REGION Network 2: Auto Initiated = Set Step to 1
   // Once the pulse has expired, with the system still in automatic, the step is set to 1
   RUNG wire#powerrail
      { S7_Templates := "SrcType := Int" } EQ_Contact(in1 := #CRNT_STEP, in2 := 0)
      I_Contact( #RST )
      Move(in := 1, out1 => #CRNT_STEP)
   END_RUNG
   // the same network as SCL:
   IF (#CRNT_STEP = 0) AND NOT #RST THEN #CRNT_STEP := 1; END_IF;
END_REGION

REGION Network 3: Sequence Running
   // Determination that the sequence is running
   RUNG wire#powerrail
      { S7_Templates := "SrcType := Int" } NE_Contact(in1 := #CRNT_STEP, in2 := 0)
      Coil( #RNG )
   END_RUNG
   // the same network as SCL:
   #RNG := #CRNT_STEP <> 0;
END_REGION

REGION Network 4: Step 001 = Confirm Auto Conditions Ok
   // Requires all conditions for auto ok to proceed
   RUNG wire#powerrail
      #STEP_001(SN := 1, CS := #CRNT_STEP, MST := "86_Times".STEP_MAX_TIME_STP_001, SC :=, BPFLT := true, AMST :=, FLT :=, ACT =>, DN =>)
      Contact( #STEP_001.DN )
      Move(in := 5, out1 => #CRNT_STEP)
   END_RUNG
   // the same network as SCL:
   #STEP_001(SN := 1, CS := #CRNT_STEP, MST := "86_Times".STEP_MAX_TIME_STP_001, BPFLT := true, ENO => #_w1);   // "500_SEQ_STEP"
   IF #_w1 AND #STEP_001.DN THEN #CRNT_STEP := 5; END_IF;
END_REGION

REGION Network 5: Step 005 = Wait For BWTS In Pre-Dwell or Dwell & ReOx
   // BWTS Active throughout
   RUNG wire#powerrail
      #STEP_005(SN := 5, CS := #CRNT_STEP, MST := "86_Times".STEP_MAX_TIME_STP_005, SC :=, BPFLT := true, AMST :=, FLT :=, ACT =>, DN =>)
      Contact( #STEP_005.DN )
      Move(in := 10, out1 => #CRNT_STEP)
   END_RUNG
   // the same network as SCL:
   #STEP_005(SN := 5, CS := #CRNT_STEP, MST := "86_Times".STEP_MAX_TIME_STP_005, BPFLT := true, ENO => #_w1);   // "500_SEQ_STEP"
   IF #_w1 AND #STEP_005.DN THEN #CRNT_STEP := 10; END_IF;
END_REGION

REGION Network 6: Step 010 = Wait For Prepare Gas Command (DeOx = Step 20, ReOx = Step 40)
   // BWTS Sends prepare gas command an hour prior to physical requirement
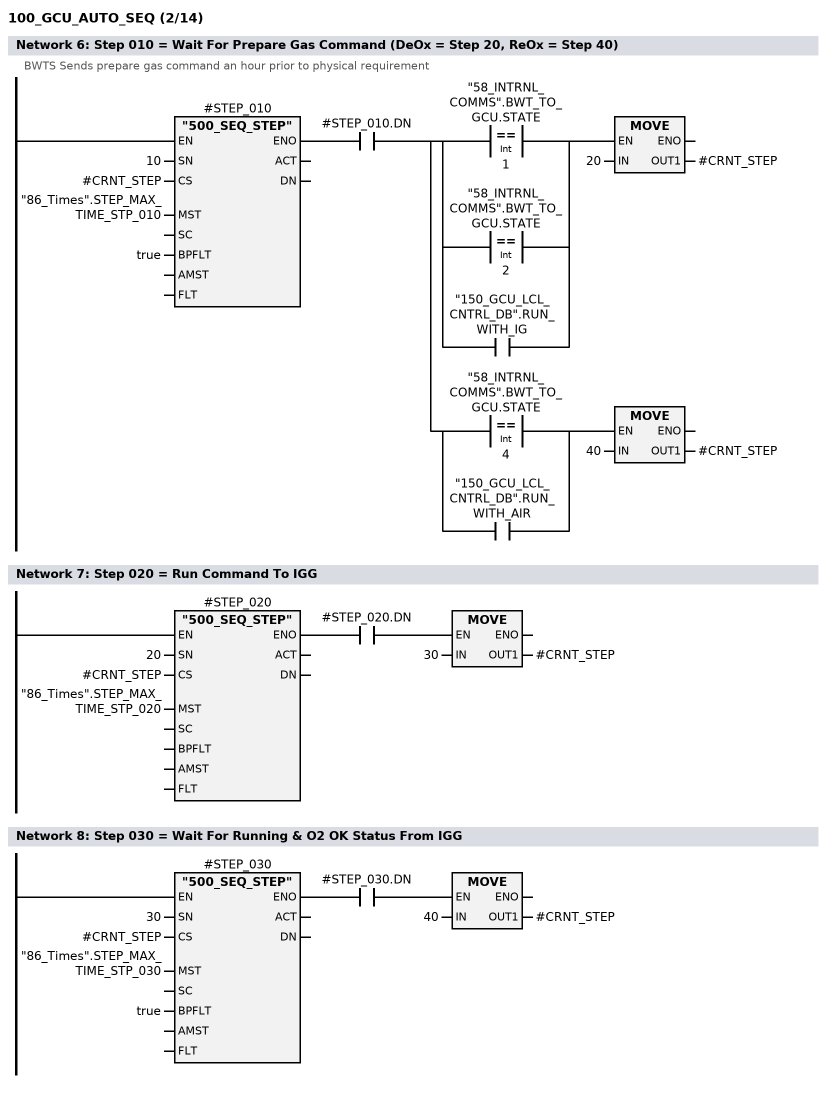
   RUNG wire#powerrail
      #STEP_010(SN := 10, CS := #CRNT_STEP, MST := "86_Times".STEP_MAX_TIME_STP_010, SC :=, BPFLT := true, AMST :=, FLT :=, ACT =>, DN =>)
      Contact( #STEP_010.DN )
      wire#w1
      { S7_Templates := "SrcType := Int" } EQ_Contact(in1 := "58_INTRNL_COMMS".BWT_TO_GCU.STATE, in2 := 1)
      wire#w2
      Move(in := 20, out1 => #CRNT_STEP)
   END_RUNG
   RUNG wire#w1
      { S7_Templates := "SrcType := Int" } EQ_Contact(in1 := "58_INTRNL_COMMS".BWT_TO_GCU.STATE, in2 := 2)
   END_RUNG wire#w2
   RUNG wire#w1
      Contact( "150_GCU_LCL_CNTRL_DB".RUN_WITH_IG )
   END_RUNG wire#w2
   RUNG wire#w1
      { S7_Templates := "SrcType := Int" } EQ_Contact(in1 := "58_INTRNL_COMMS".BWT_TO_GCU.STATE, in2 := 4)
      wire#w3
      Move(in := 40, out1 => #CRNT_STEP)
   END_RUNG
   RUNG wire#w1
      Contact( "150_GCU_LCL_CNTRL_DB".RUN_WITH_AIR )
   END_RUNG wire#w3
   // the same network as SCL:
   #STEP_010(SN := 10, CS := #CRNT_STEP, MST := "86_Times".STEP_MAX_TIME_STP_010, BPFLT := true, ENO => #_w1);   // "500_SEQ_STEP"
   #_w2 := #_w1 AND #STEP_010.DN;
   IF #_w2 AND (("58_INTRNL_COMMS".BWT_TO_GCU.STATE = 1) OR ("58_INTRNL_COMMS".BWT_TO_GCU.STATE = 2) OR "150_GCU_LCL_CNTRL_DB".RUN_WITH_IG) THEN
       #CRNT_STEP := 20;
   END_IF;
   IF #_w2 AND (("58_INTRNL_COMMS".BWT_TO_GCU.STATE = 4) OR "150_GCU_LCL_CNTRL_DB".RUN_WITH_AIR) THEN
       #CRNT_STEP := 40;
   END_IF;
END_REGION

REGION Network 7: Step 020 = Run Command To IGG
   RUNG wire#powerrail
      #STEP_020(SN := 20, CS := #CRNT_STEP, MST := "86_Times".STEP_MAX_TIME_STP_020, SC :=, BPFLT :=, AMST :=, FLT :=, ACT =>, DN =>)
      Contact( #STEP_020.DN )
      Move(in := 30, out1 => #CRNT_STEP)
   END_RUNG
   // the same network as SCL:
   #STEP_020(SN := 20, CS := #CRNT_STEP, MST := "86_Times".STEP_MAX_TIME_STP_020, ENO => #_w1);   // "500_SEQ_STEP"
   IF #_w1 AND #STEP_020.DN THEN #CRNT_STEP := 30; END_IF;
END_REGION

REGION Network 8: Step 030 = Wait For Running & O2 OK Status From IGG
   RUNG wire#powerrail
      #STEP_030(SN := 30, CS := #CRNT_STEP, MST := "86_Times".STEP_MAX_TIME_STP_030, SC :=, BPFLT := true, AMST :=, FLT :=, ACT =>, DN =>)
      Contact( #STEP_030.DN )
      Move(in := 40, out1 => #CRNT_STEP)
   END_RUNG
   // the same network as SCL:
   #STEP_030(SN := 30, CS := #CRNT_STEP, MST := "86_Times".STEP_MAX_TIME_STP_030, BPFLT := true, ENO => #_w1);   // "500_SEQ_STEP"
   IF #_w1 AND #STEP_030.DN THEN #CRNT_STEP := 40; END_IF;
END_REGION

REGION Network 9: Step 040 = Wait For Supply Gas Command
   // Gas available status to BWTS
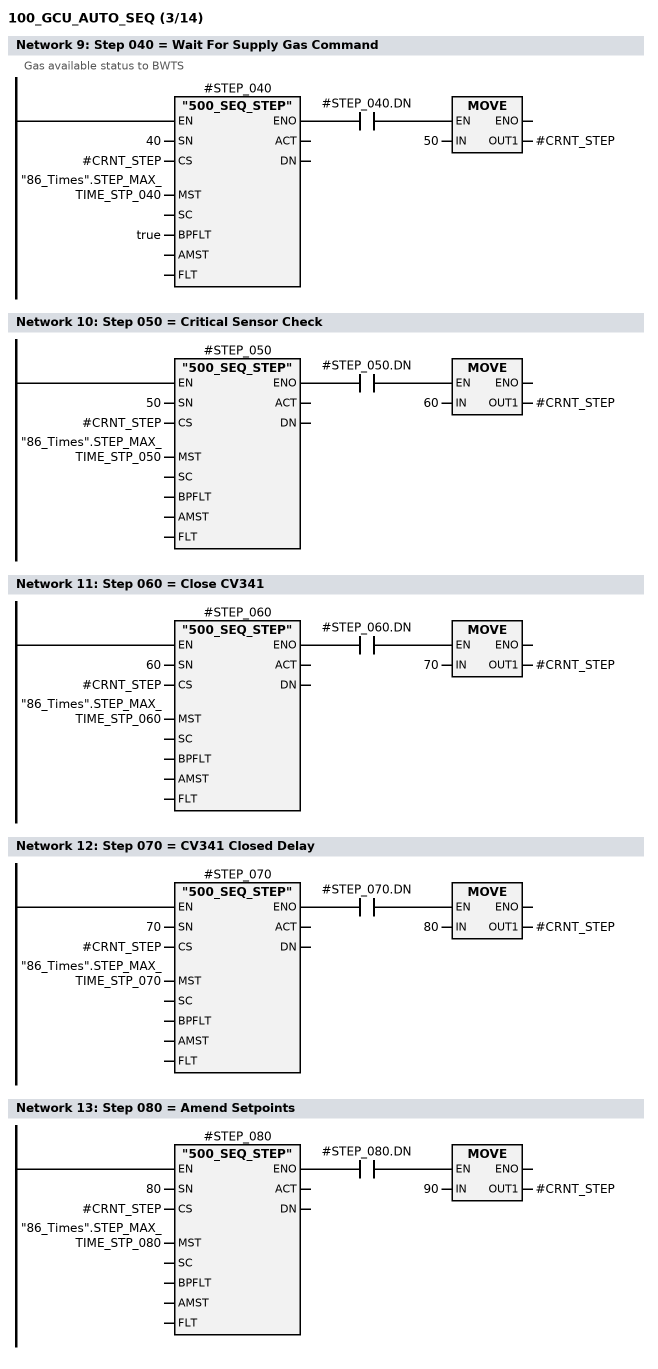
   RUNG wire#powerrail
      #STEP_040(SN := 40, CS := #CRNT_STEP, MST := "86_Times".STEP_MAX_TIME_STP_040, SC :=, BPFLT := true, AMST :=, FLT :=, ACT =>, DN =>)
      Contact( #STEP_040.DN )
      Move(in := 50, out1 => #CRNT_STEP)
   END_RUNG
   // the same network as SCL:
   #STEP_040(SN := 40, CS := #CRNT_STEP, MST := "86_Times".STEP_MAX_TIME_STP_040, BPFLT := true, ENO => #_w1);   // "500_SEQ_STEP"
   IF #_w1 AND #STEP_040.DN THEN #CRNT_STEP := 50; END_IF;
END_REGION

REGION Network 10: Step 050 = Critical Sensor Check
   RUNG wire#powerrail
      #STEP_050(SN := 50, CS := #CRNT_STEP, MST := "86_Times".STEP_MAX_TIME_STP_050, SC :=, BPFLT :=, AMST :=, FLT :=, ACT =>, DN =>)
      Contact( #STEP_050.DN )
      Move(in := 60, out1 => #CRNT_STEP)
   END_RUNG
   // the same network as SCL:
   #STEP_050(SN := 50, CS := #CRNT_STEP, MST := "86_Times".STEP_MAX_TIME_STP_050, ENO => #_w1);   // "500_SEQ_STEP"
   IF #_w1 AND #STEP_050.DN THEN #CRNT_STEP := 60; END_IF;
END_REGION

REGION Network 11: Step 060 = Close CV341
   RUNG wire#powerrail
      #STEP_060(SN := 60, CS := #CRNT_STEP, MST := "86_Times".STEP_MAX_TIME_STP_060, SC :=, BPFLT :=, AMST :=, FLT :=, ACT =>, DN =>)
      Contact( #STEP_060.DN )
      Move(in := 70, out1 => #CRNT_STEP)
   END_RUNG
   // the same network as SCL:
   #STEP_060(SN := 60, CS := #CRNT_STEP, MST := "86_Times".STEP_MAX_TIME_STP_060, ENO => #_w1);   // "500_SEQ_STEP"
   IF #_w1 AND #STEP_060.DN THEN #CRNT_STEP := 70; END_IF;
END_REGION

REGION Network 12: Step 070 = CV341 Closed Delay
   RUNG wire#powerrail
      #STEP_070(SN := 70, CS := #CRNT_STEP, MST := "86_Times".STEP_MAX_TIME_STP_070, SC :=, BPFLT :=, AMST :=, FLT :=, ACT =>, DN =>)
      Contact( #STEP_070.DN )
      Move(in := 80, out1 => #CRNT_STEP)
   END_RUNG
   // the same network as SCL:
   #STEP_070(SN := 70, CS := #CRNT_STEP, MST := "86_Times".STEP_MAX_TIME_STP_070, ENO => #_w1);   // "500_SEQ_STEP"
   IF #_w1 AND #STEP_070.DN THEN #CRNT_STEP := 80; END_IF;
END_REGION

REGION Network 13: Step 080 = Amend Setpoints
   RUNG wire#powerrail
      #STEP_080(SN := 80, CS := #CRNT_STEP, MST := "86_Times".STEP_MAX_TIME_STP_080, SC :=, BPFLT :=, AMST :=, FLT :=, ACT =>, DN =>)
      Contact( #STEP_080.DN )
      Move(in := 90, out1 => #CRNT_STEP)
   END_RUNG
   // the same network as SCL:
   #STEP_080(SN := 80, CS := #CRNT_STEP, MST := "86_Times".STEP_MAX_TIME_STP_080, ENO => #_w1);   // "500_SEQ_STEP"
   IF #_w1 AND #STEP_080.DN THEN #CRNT_STEP := 90; END_IF;
END_REGION

REGION Network 14: Step 090 = Open CV358
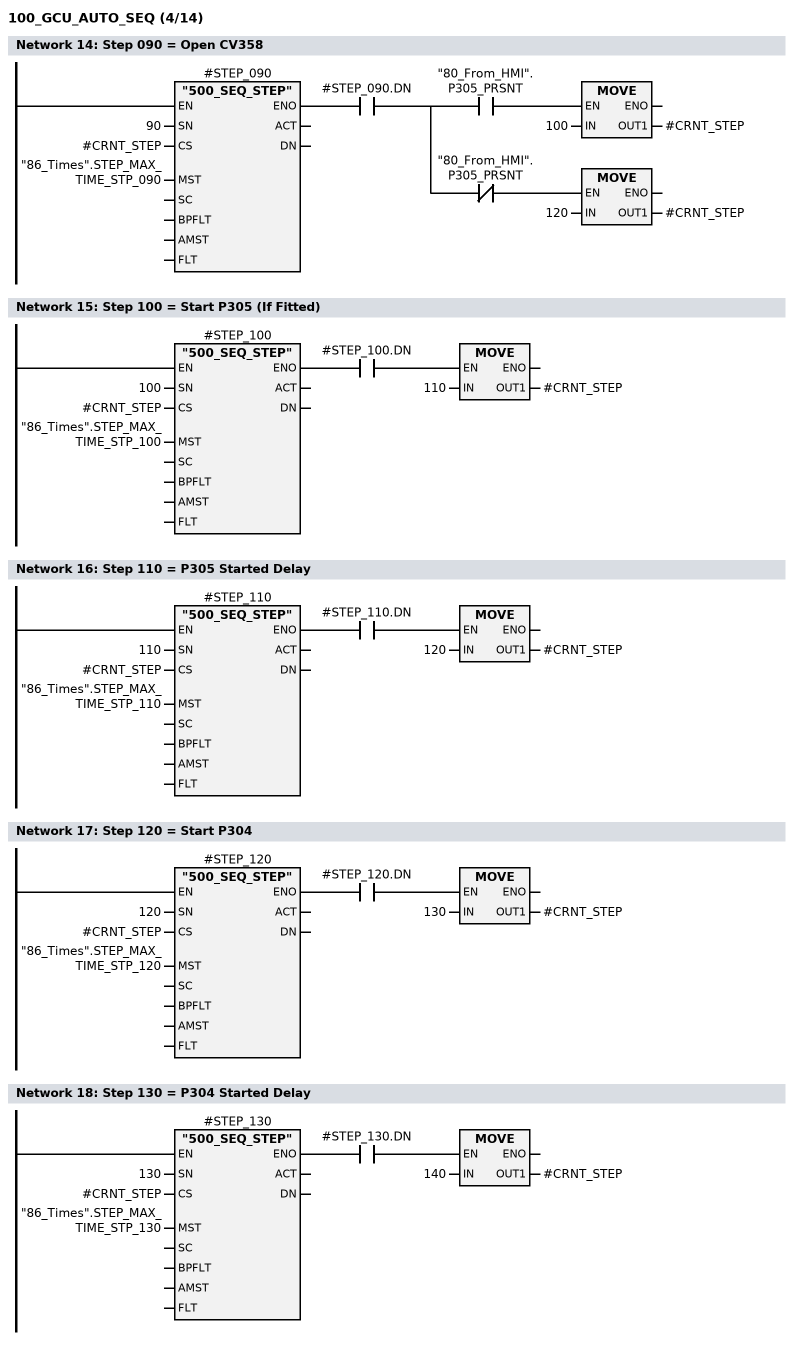
   RUNG wire#powerrail
      #STEP_090(SN := 90, CS := #CRNT_STEP, MST := "86_Times".STEP_MAX_TIME_STP_090, SC :=, BPFLT :=, AMST :=, FLT :=, ACT =>, DN =>)
      Contact( #STEP_090.DN )
      wire#w1
      Contact( "80_From_HMI".P305_PRSNT )
      Move(in := 100, out1 => #CRNT_STEP)
   END_RUNG
   RUNG wire#w1
      I_Contact( "80_From_HMI".P305_PRSNT )
      Move(in := 120, out1 => #CRNT_STEP)
   END_RUNG
   // the same network as SCL:
   #STEP_090(SN := 90, CS := #CRNT_STEP, MST := "86_Times".STEP_MAX_TIME_STP_090, ENO => #_w1);   // "500_SEQ_STEP"
   #_w2 := #_w1 AND #STEP_090.DN;
   IF #_w2 AND "80_From_HMI".P305_PRSNT THEN #CRNT_STEP := 100; END_IF;
   IF #_w2 AND NOT "80_From_HMI".P305_PRSNT THEN #CRNT_STEP := 120; END_IF;
END_REGION

REGION Network 15: Step 100 = Start P305 (If Fitted)
   RUNG wire#powerrail
      #STEP_100(SN := 100, CS := #CRNT_STEP, MST := "86_Times".STEP_MAX_TIME_STP_100, SC :=, BPFLT :=, AMST :=, FLT :=, ACT =>, DN =>)
      Contact( #STEP_100.DN )
      Move(in := 110, out1 => #CRNT_STEP)
   END_RUNG
   // the same network as SCL:
   #STEP_100(SN := 100, CS := #CRNT_STEP, MST := "86_Times".STEP_MAX_TIME_STP_100, ENO => #_w1);   // "500_SEQ_STEP"
   IF #_w1 AND #STEP_100.DN THEN #CRNT_STEP := 110; END_IF;
END_REGION

REGION Network 16: Step 110 = P305 Started Delay
   RUNG wire#powerrail
      #STEP_110(SN := 110, CS := #CRNT_STEP, MST := "86_Times".STEP_MAX_TIME_STP_110, SC :=, BPFLT :=, AMST :=, FLT :=, ACT =>, DN =>)
      Contact( #STEP_110.DN )
      Move(in := 120, out1 => #CRNT_STEP)
   END_RUNG
   // the same network as SCL:
   #STEP_110(SN := 110, CS := #CRNT_STEP, MST := "86_Times".STEP_MAX_TIME_STP_110, ENO => #_w1);   // "500_SEQ_STEP"
   IF #_w1 AND #STEP_110.DN THEN #CRNT_STEP := 120; END_IF;
END_REGION

REGION Network 17: Step 120 = Start P304
   RUNG wire#powerrail
      #STEP_120(SN := 120, CS := #CRNT_STEP, MST := "86_Times".STEP_MAX_TIME_STP_120, SC :=, BPFLT :=, AMST :=, FLT :=, ACT =>, DN =>)
      Contact( #STEP_120.DN )
      Move(in := 130, out1 => #CRNT_STEP)
   END_RUNG
   // the same network as SCL:
   #STEP_120(SN := 120, CS := #CRNT_STEP, MST := "86_Times".STEP_MAX_TIME_STP_120, ENO => #_w1);   // "500_SEQ_STEP"
   IF #_w1 AND #STEP_120.DN THEN #CRNT_STEP := 130; END_IF;
END_REGION

REGION Network 18: Step 130 = P304 Started Delay
   RUNG wire#powerrail
      #STEP_130(SN := 130, CS := #CRNT_STEP, MST := "86_Times".STEP_MAX_TIME_STP_130, SC :=, BPFLT :=, AMST :=, FLT :=, ACT =>, DN =>)
      Contact( #STEP_130.DN )
      Move(in := 140, out1 => #CRNT_STEP)
   END_RUNG
   // the same network as SCL:
   #STEP_130(SN := 130, CS := #CRNT_STEP, MST := "86_Times".STEP_MAX_TIME_STP_130, ENO => #_w1);   // "500_SEQ_STEP"
   IF #_w1 AND #STEP_130.DN THEN #CRNT_STEP := 140; END_IF;
END_REGION

REGION Network 19: Step 140 = GCU Tank Pre-Fill Delay
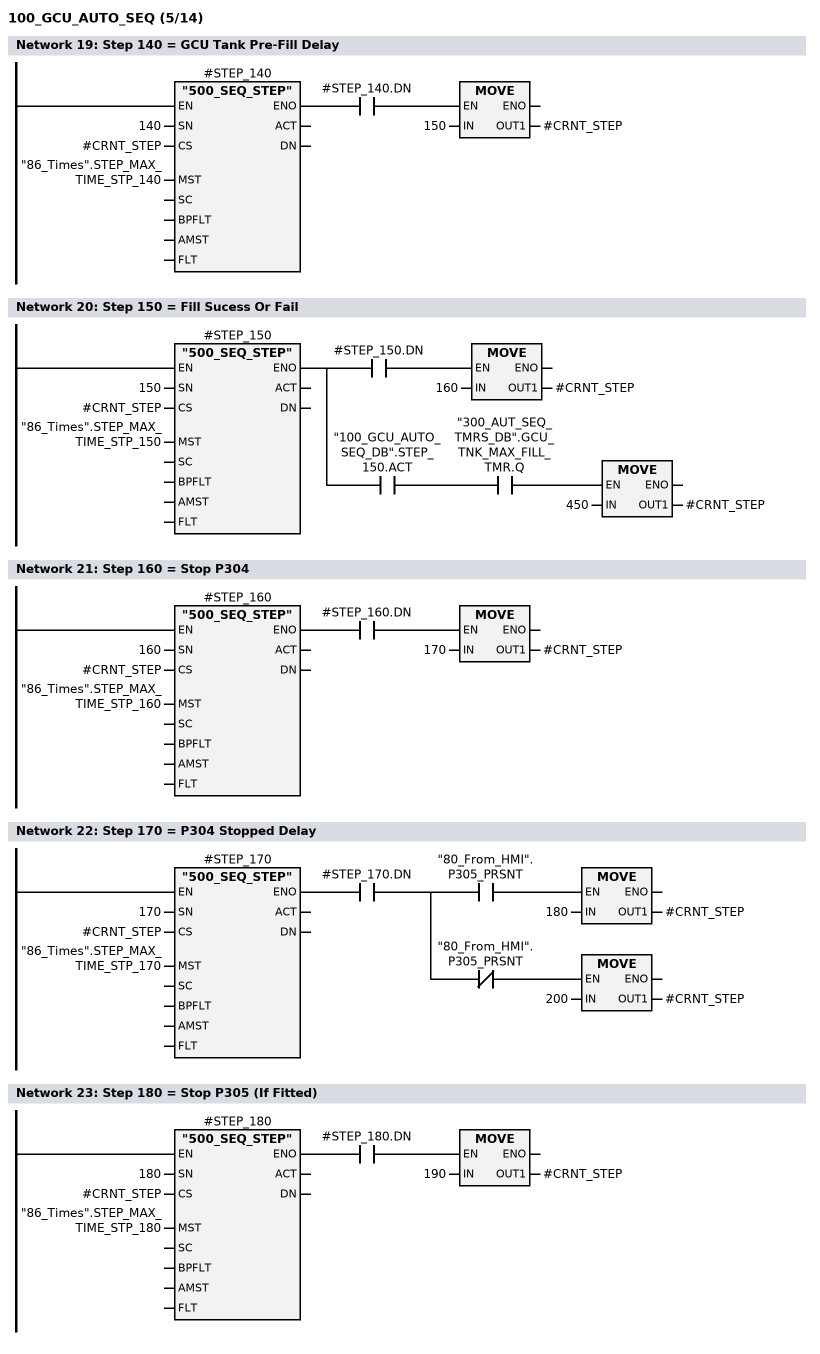
   RUNG wire#powerrail
      #STEP_140(SN := 140, CS := #CRNT_STEP, MST := "86_Times".STEP_MAX_TIME_STP_140, SC :=, BPFLT :=, AMST :=, FLT :=, ACT =>, DN =>)
      Contact( #STEP_140.DN )
      Move(in := 150, out1 => #CRNT_STEP)
   END_RUNG
   // the same network as SCL:
   #STEP_140(SN := 140, CS := #CRNT_STEP, MST := "86_Times".STEP_MAX_TIME_STP_140, ENO => #_w1);   // "500_SEQ_STEP"
   IF #_w1 AND #STEP_140.DN THEN #CRNT_STEP := 150; END_IF;
END_REGION

REGION Network 20: Step 150 = Fill Sucess Or Fail
   RUNG wire#powerrail
      #STEP_150(SN := 150, CS := #CRNT_STEP, MST := "86_Times".STEP_MAX_TIME_STP_150, SC :=, BPFLT :=, AMST :=, FLT :=, ACT =>, DN =>)
      wire#w1
      Contact( #STEP_150.DN )
      Move(in := 160, out1 => #CRNT_STEP)
   END_RUNG
   RUNG wire#w1
      Contact( "100_GCU_AUTO_SEQ_DB".STEP_150.ACT )
      Contact( "300_AUT_SEQ_TMRS_DB".GCU_TNK_MAX_FILL_TMR.Q )
      Move(in := 450, out1 => #CRNT_STEP)
   END_RUNG
   // the same network as SCL:
   #STEP_150(SN := 150, CS := #CRNT_STEP, MST := "86_Times".STEP_MAX_TIME_STP_150, ENO => #_w1);   // "500_SEQ_STEP"
   IF #_w1 AND #STEP_150.DN THEN #CRNT_STEP := 160; END_IF;
   IF #_w1 AND "100_GCU_AUTO_SEQ_DB".STEP_150.ACT AND "300_AUT_SEQ_TMRS_DB".GCU_TNK_MAX_FILL_TMR.Q THEN
       #CRNT_STEP := 450;
   END_IF;
END_REGION

REGION Network 21: Step 160 = Stop P304
   RUNG wire#powerrail
      #STEP_160(SN := 160, CS := #CRNT_STEP, MST := "86_Times".STEP_MAX_TIME_STP_160, SC :=, BPFLT :=, AMST :=, FLT :=, ACT =>, DN =>)
      Contact( #STEP_160.DN )
      Move(in := 170, out1 => #CRNT_STEP)
   END_RUNG
   // the same network as SCL:
   #STEP_160(SN := 160, CS := #CRNT_STEP, MST := "86_Times".STEP_MAX_TIME_STP_160, ENO => #_w1);   // "500_SEQ_STEP"
   IF #_w1 AND #STEP_160.DN THEN #CRNT_STEP := 170; END_IF;
END_REGION

REGION Network 22: Step 170 = P304 Stopped Delay
   RUNG wire#powerrail
      #STEP_170(SN := 170, CS := #CRNT_STEP, MST := "86_Times".STEP_MAX_TIME_STP_170, SC :=, BPFLT :=, AMST :=, FLT :=, ACT =>, DN =>)
      Contact( #STEP_170.DN )
      wire#w1
      Contact( "80_From_HMI".P305_PRSNT )
      Move(in := 180, out1 => #CRNT_STEP)
   END_RUNG
   RUNG wire#w1
      I_Contact( "80_From_HMI".P305_PRSNT )
      Move(in := 200, out1 => #CRNT_STEP)
   END_RUNG
   // the same network as SCL:
   #STEP_170(SN := 170, CS := #CRNT_STEP, MST := "86_Times".STEP_MAX_TIME_STP_170, ENO => #_w1);   // "500_SEQ_STEP"
   #_w2 := #_w1 AND #STEP_170.DN;
   IF #_w2 AND "80_From_HMI".P305_PRSNT THEN #CRNT_STEP := 180; END_IF;
   IF #_w2 AND NOT "80_From_HMI".P305_PRSNT THEN #CRNT_STEP := 200; END_IF;
END_REGION

REGION Network 23: Step 180 = Stop P305 (If Fitted)
   RUNG wire#powerrail
      #STEP_180(SN := 180, CS := #CRNT_STEP, MST := "86_Times".STEP_MAX_TIME_STP_180, SC :=, BPFLT :=, AMST :=, FLT :=, ACT =>, DN =>)
      Contact( #STEP_180.DN )
      Move(in := 190, out1 => #CRNT_STEP)
   END_RUNG
   // the same network as SCL:
   #STEP_180(SN := 180, CS := #CRNT_STEP, MST := "86_Times".STEP_MAX_TIME_STP_180, ENO => #_w1);   // "500_SEQ_STEP"
   IF #_w1 AND #STEP_180.DN THEN #CRNT_STEP := 190; END_IF;
END_REGION

REGION Network 24: Step 190 = P305 Stopped Delay
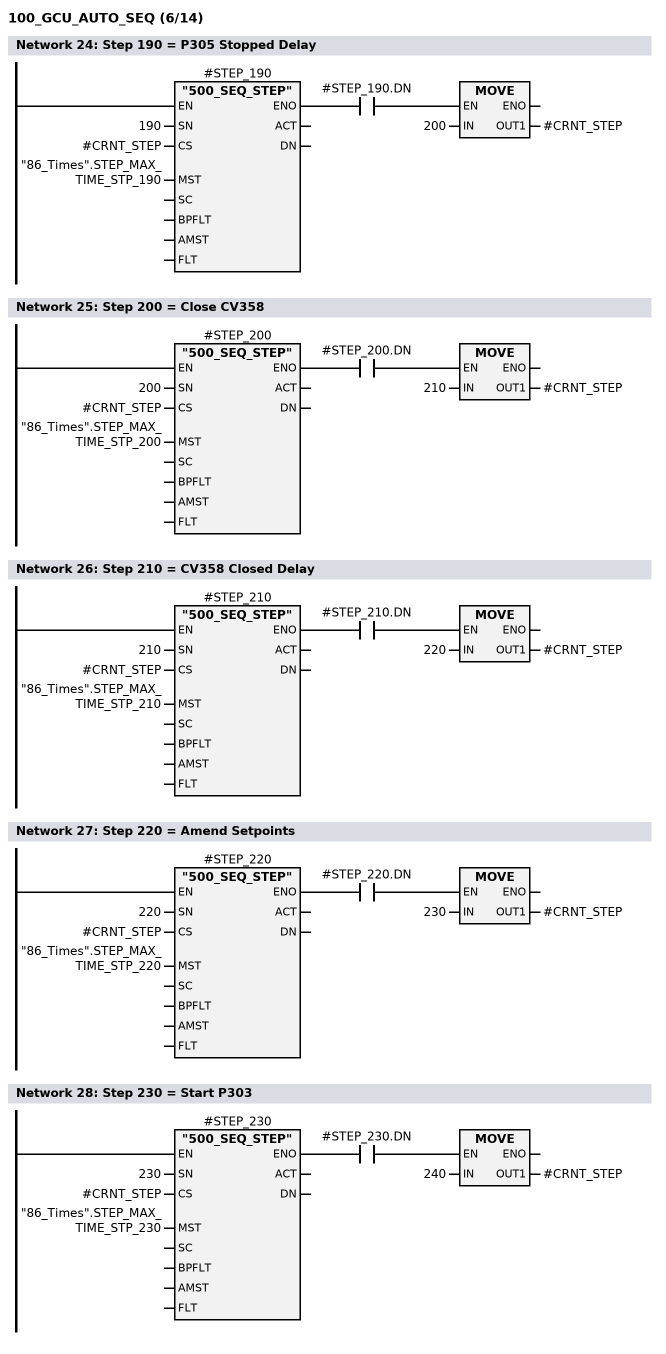
   RUNG wire#powerrail
      #STEP_190(SN := 190, CS := #CRNT_STEP, MST := "86_Times".STEP_MAX_TIME_STP_190, SC :=, BPFLT :=, AMST :=, FLT :=, ACT =>, DN =>)
      Contact( #STEP_190.DN )
      Move(in := 200, out1 => #CRNT_STEP)
   END_RUNG
   // the same network as SCL:
   #STEP_190(SN := 190, CS := #CRNT_STEP, MST := "86_Times".STEP_MAX_TIME_STP_190, ENO => #_w1);   // "500_SEQ_STEP"
   IF #_w1 AND #STEP_190.DN THEN #CRNT_STEP := 200; END_IF;
END_REGION

REGION Network 25: Step 200 = Close CV358
   RUNG wire#powerrail
      #STEP_200(SN := 200, CS := #CRNT_STEP, MST := "86_Times".STEP_MAX_TIME_STP_200, SC :=, BPFLT :=, AMST :=, FLT :=, ACT =>, DN =>)
      Contact( #STEP_200.DN )
      Move(in := 210, out1 => #CRNT_STEP)
   END_RUNG
   // the same network as SCL:
   #STEP_200(SN := 200, CS := #CRNT_STEP, MST := "86_Times".STEP_MAX_TIME_STP_200, ENO => #_w1);   // "500_SEQ_STEP"
   IF #_w1 AND #STEP_200.DN THEN #CRNT_STEP := 210; END_IF;
END_REGION

REGION Network 26: Step 210 = CV358 Closed Delay
   RUNG wire#powerrail
      #STEP_210(SN := 210, CS := #CRNT_STEP, MST := "86_Times".STEP_MAX_TIME_STP_210, SC :=, BPFLT :=, AMST :=, FLT :=, ACT =>, DN =>)
      Contact( #STEP_210.DN )
      Move(in := 220, out1 => #CRNT_STEP)
   END_RUNG
   // the same network as SCL:
   #STEP_210(SN := 210, CS := #CRNT_STEP, MST := "86_Times".STEP_MAX_TIME_STP_210, ENO => #_w1);   // "500_SEQ_STEP"
   IF #_w1 AND #STEP_210.DN THEN #CRNT_STEP := 220; END_IF;
END_REGION

REGION Network 27: Step 220 = Amend Setpoints
   RUNG wire#powerrail
      #STEP_220(SN := 220, CS := #CRNT_STEP, MST := "86_Times".STEP_MAX_TIME_STP_220, SC :=, BPFLT :=, AMST :=, FLT :=, ACT =>, DN =>)
      Contact( #STEP_220.DN )
      Move(in := 230, out1 => #CRNT_STEP)
   END_RUNG
   // the same network as SCL:
   #STEP_220(SN := 220, CS := #CRNT_STEP, MST := "86_Times".STEP_MAX_TIME_STP_220, ENO => #_w1);   // "500_SEQ_STEP"
   IF #_w1 AND #STEP_220.DN THEN #CRNT_STEP := 230; END_IF;
END_REGION

REGION Network 28: Step 230 = Start P303
   RUNG wire#powerrail
      #STEP_230(SN := 230, CS := #CRNT_STEP, MST := "86_Times".STEP_MAX_TIME_STP_230, SC :=, BPFLT :=, AMST :=, FLT :=, ACT =>, DN =>)
      Contact( #STEP_230.DN )
      Move(in := 240, out1 => #CRNT_STEP)
   END_RUNG
   // the same network as SCL:
   #STEP_230(SN := 230, CS := #CRNT_STEP, MST := "86_Times".STEP_MAX_TIME_STP_230, ENO => #_w1);   // "500_SEQ_STEP"
   IF #_w1 AND #STEP_230.DN THEN #CRNT_STEP := 240; END_IF;
END_REGION

REGION Network 29: Step 240 = P303 Started Delay
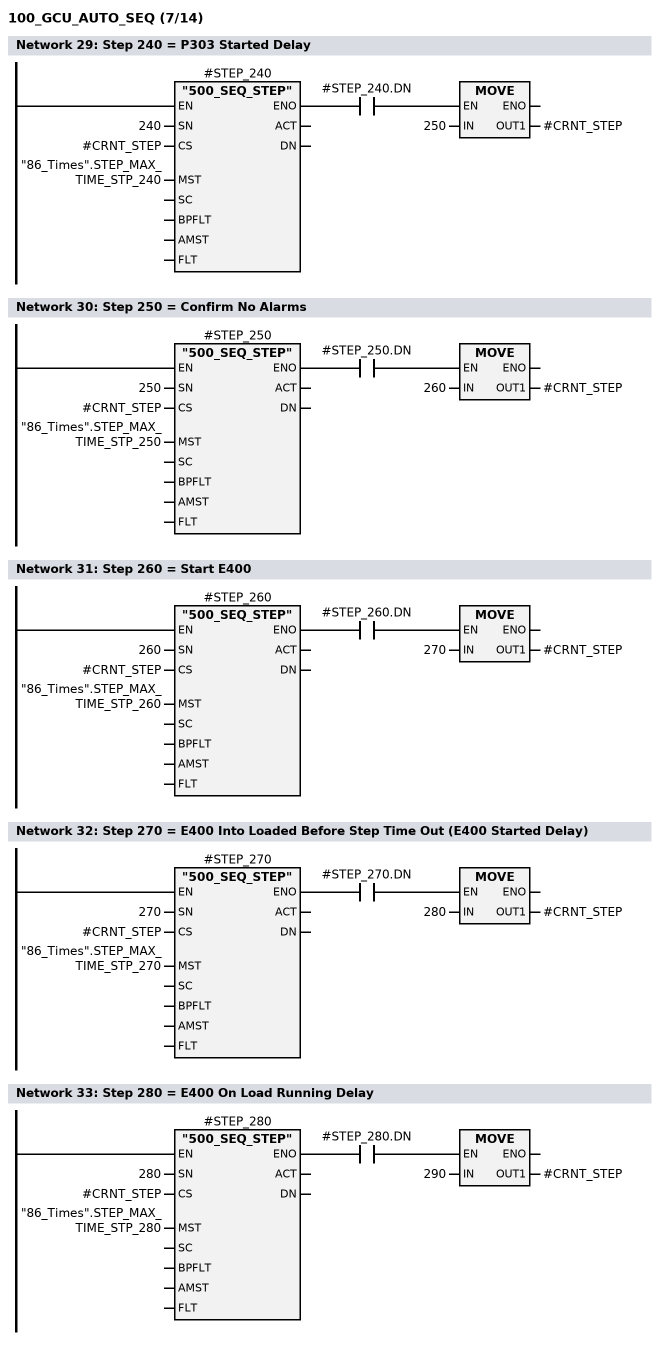
   RUNG wire#powerrail
      #STEP_240(SN := 240, CS := #CRNT_STEP, MST := "86_Times".STEP_MAX_TIME_STP_240, SC :=, BPFLT :=, AMST :=, FLT :=, ACT =>, DN =>)
      Contact( #STEP_240.DN )
      Move(in := 250, out1 => #CRNT_STEP)
   END_RUNG
   // the same network as SCL:
   #STEP_240(SN := 240, CS := #CRNT_STEP, MST := "86_Times".STEP_MAX_TIME_STP_240, ENO => #_w1);   // "500_SEQ_STEP"
   IF #_w1 AND #STEP_240.DN THEN #CRNT_STEP := 250; END_IF;
END_REGION

REGION Network 30: Step 250 = Confirm No Alarms
   RUNG wire#powerrail
      #STEP_250(SN := 250, CS := #CRNT_STEP, MST := "86_Times".STEP_MAX_TIME_STP_250, SC :=, BPFLT :=, AMST :=, FLT :=, ACT =>, DN =>)
      Contact( #STEP_250.DN )
      Move(in := 260, out1 => #CRNT_STEP)
   END_RUNG
   // the same network as SCL:
   #STEP_250(SN := 250, CS := #CRNT_STEP, MST := "86_Times".STEP_MAX_TIME_STP_250, ENO => #_w1);   // "500_SEQ_STEP"
   IF #_w1 AND #STEP_250.DN THEN #CRNT_STEP := 260; END_IF;
END_REGION

REGION Network 31: Step 260 = Start E400
   RUNG wire#powerrail
      #STEP_260(SN := 260, CS := #CRNT_STEP, MST := "86_Times".STEP_MAX_TIME_STP_260, SC :=, BPFLT :=, AMST :=, FLT :=, ACT =>, DN =>)
      Contact( #STEP_260.DN )
      Move(in := 270, out1 => #CRNT_STEP)
   END_RUNG
   // the same network as SCL:
   #STEP_260(SN := 260, CS := #CRNT_STEP, MST := "86_Times".STEP_MAX_TIME_STP_260, ENO => #_w1);   // "500_SEQ_STEP"
   IF #_w1 AND #STEP_260.DN THEN #CRNT_STEP := 270; END_IF;
END_REGION

REGION Network 32: Step 270 = E400 Into Loaded Before Step Time Out (E400 Started Delay)
   RUNG wire#powerrail
      #STEP_270(SN := 270, CS := #CRNT_STEP, MST := "86_Times".STEP_MAX_TIME_STP_270, SC :=, BPFLT :=, AMST :=, FLT :=, ACT =>, DN =>)
      Contact( #STEP_270.DN )
      Move(in := 280, out1 => #CRNT_STEP)
   END_RUNG
   // the same network as SCL:
   #STEP_270(SN := 270, CS := #CRNT_STEP, MST := "86_Times".STEP_MAX_TIME_STP_270, ENO => #_w1);   // "500_SEQ_STEP"
   IF #_w1 AND #STEP_270.DN THEN #CRNT_STEP := 280; END_IF;
END_REGION

REGION Network 33: Step 280 = E400 On Load Running Delay
   RUNG wire#powerrail
      #STEP_280(SN := 280, CS := #CRNT_STEP, MST := "86_Times".STEP_MAX_TIME_STP_280, SC :=, BPFLT :=, AMST :=, FLT :=, ACT =>, DN =>)
      Contact( #STEP_280.DN )
      Move(in := 290, out1 => #CRNT_STEP)
   END_RUNG
   // the same network as SCL:
   #STEP_280(SN := 280, CS := #CRNT_STEP, MST := "86_Times".STEP_MAX_TIME_STP_280, ENO => #_w1);   // "500_SEQ_STEP"
   IF #_w1 AND #STEP_280.DN THEN #CRNT_STEP := 290; END_IF;
END_REGION

REGION Network 34: Step 290 = CV405 Modulation Start & PIT416 Target Ramp Run
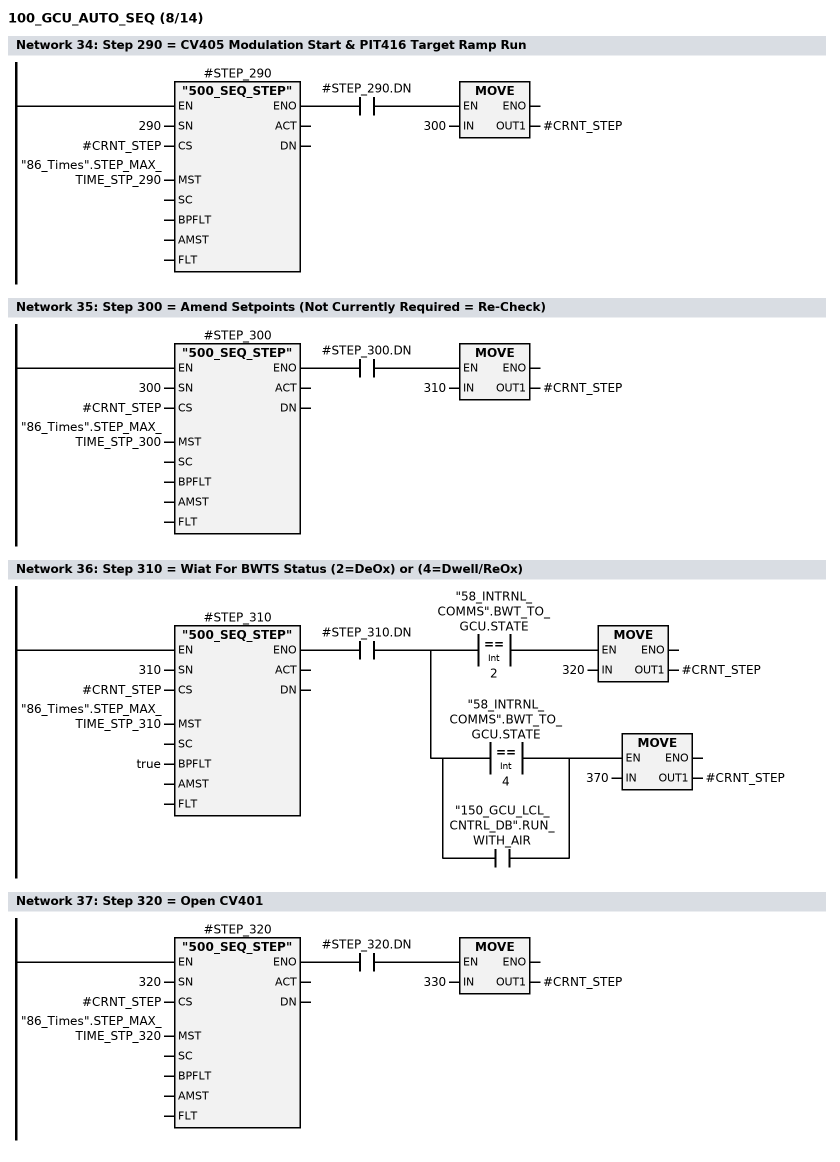
   RUNG wire#powerrail
      #STEP_290(SN := 290, CS := #CRNT_STEP, MST := "86_Times".STEP_MAX_TIME_STP_290, SC :=, BPFLT :=, AMST :=, FLT :=, ACT =>, DN =>)
      Contact( #STEP_290.DN )
      Move(in := 300, out1 => #CRNT_STEP)
   END_RUNG
   // the same network as SCL:
   #STEP_290(SN := 290, CS := #CRNT_STEP, MST := "86_Times".STEP_MAX_TIME_STP_290, ENO => #_w1);   // "500_SEQ_STEP"
   IF #_w1 AND #STEP_290.DN THEN #CRNT_STEP := 300; END_IF;
END_REGION

REGION Network 35: Step 300 = Amend Setpoints (Not Currently Required = Re-Check)
   RUNG wire#powerrail
      #STEP_300(SN := 300, CS := #CRNT_STEP, MST := "86_Times".STEP_MAX_TIME_STP_300, SC :=, BPFLT :=, AMST :=, FLT :=, ACT =>, DN =>)
      Contact( #STEP_300.DN )
      Move(in := 310, out1 => #CRNT_STEP)
   END_RUNG
   // the same network as SCL:
   #STEP_300(SN := 300, CS := #CRNT_STEP, MST := "86_Times".STEP_MAX_TIME_STP_300, ENO => #_w1);   // "500_SEQ_STEP"
   IF #_w1 AND #STEP_300.DN THEN #CRNT_STEP := 310; END_IF;
END_REGION

REGION Network 36: Step 310 = Wiat For BWTS Status (2=DeOx) or (4=Dwell/ReOx)
   RUNG wire#powerrail
      #STEP_310(SN := 310, CS := #CRNT_STEP, MST := "86_Times".STEP_MAX_TIME_STP_310, SC :=, BPFLT := true, AMST :=, FLT :=, ACT =>, DN =>)
      Contact( #STEP_310.DN )
      wire#w1
      { S7_Templates := "SrcType := Int" } EQ_Contact(in1 := "58_INTRNL_COMMS".BWT_TO_GCU.STATE, in2 := 2)
      Move(in := 320, out1 => #CRNT_STEP)
   END_RUNG
   RUNG wire#w1
      { S7_Templates := "SrcType := Int" } EQ_Contact(in1 := "58_INTRNL_COMMS".BWT_TO_GCU.STATE, in2 := 4)
      wire#w2
      Move(in := 370, out1 => #CRNT_STEP)
   END_RUNG
   RUNG wire#w1
      Contact( "150_GCU_LCL_CNTRL_DB".RUN_WITH_AIR )
   END_RUNG wire#w2
   // the same network as SCL:
   #STEP_310(SN := 310, CS := #CRNT_STEP, MST := "86_Times".STEP_MAX_TIME_STP_310, BPFLT := true, ENO => #_w1);   // "500_SEQ_STEP"
   #_w2 := #_w1 AND #STEP_310.DN;
   IF #_w2 AND ("58_INTRNL_COMMS".BWT_TO_GCU.STATE = 2) THEN #CRNT_STEP := 320; END_IF;
   IF #_w2 AND (("58_INTRNL_COMMS".BWT_TO_GCU.STATE = 4) OR "150_GCU_LCL_CNTRL_DB".RUN_WITH_AIR) THEN
       #CRNT_STEP := 370;
   END_IF;
END_REGION

REGION Network 37: Step 320 = Open CV401
   RUNG wire#powerrail
      #STEP_320(SN := 320, CS := #CRNT_STEP, MST := "86_Times".STEP_MAX_TIME_STP_320, SC :=, BPFLT :=, AMST :=, FLT :=, ACT =>, DN =>)
      Contact( #STEP_320.DN )
      Move(in := 330, out1 => #CRNT_STEP)
   END_RUNG
   // the same network as SCL:
   #STEP_320(SN := 320, CS := #CRNT_STEP, MST := "86_Times".STEP_MAX_TIME_STP_320, ENO => #_w1);   // "500_SEQ_STEP"
   IF #_w1 AND #STEP_320.DN THEN #CRNT_STEP := 330; END_IF;
END_REGION

REGION Network 38: Step 330 = CV401 Opened Delay
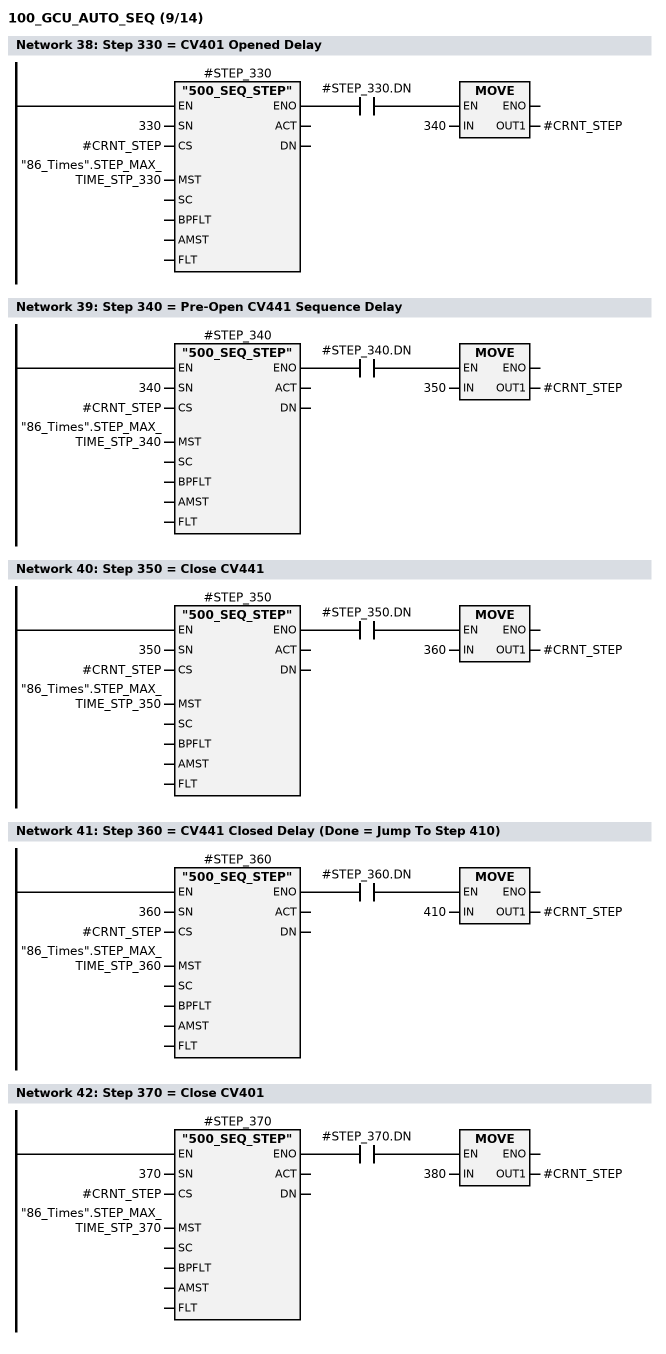
   RUNG wire#powerrail
      #STEP_330(SN := 330, CS := #CRNT_STEP, MST := "86_Times".STEP_MAX_TIME_STP_330, SC :=, BPFLT :=, AMST :=, FLT :=, ACT =>, DN =>)
      Contact( #STEP_330.DN )
      Move(in := 340, out1 => #CRNT_STEP)
   END_RUNG
   // the same network as SCL:
   #STEP_330(SN := 330, CS := #CRNT_STEP, MST := "86_Times".STEP_MAX_TIME_STP_330, ENO => #_w1);   // "500_SEQ_STEP"
   IF #_w1 AND #STEP_330.DN THEN #CRNT_STEP := 340; END_IF;
END_REGION

REGION Network 39: Step 340 = Pre-Open CV441 Sequence Delay
   RUNG wire#powerrail
      #STEP_340(SN := 340, CS := #CRNT_STEP, MST := "86_Times".STEP_MAX_TIME_STP_340, SC :=, BPFLT :=, AMST :=, FLT :=, ACT =>, DN =>)
      Contact( #STEP_340.DN )
      Move(in := 350, out1 => #CRNT_STEP)
   END_RUNG
   // the same network as SCL:
   #STEP_340(SN := 340, CS := #CRNT_STEP, MST := "86_Times".STEP_MAX_TIME_STP_340, ENO => #_w1);   // "500_SEQ_STEP"
   IF #_w1 AND #STEP_340.DN THEN #CRNT_STEP := 350; END_IF;
END_REGION

REGION Network 40: Step 350 = Close CV441
   RUNG wire#powerrail
      #STEP_350(SN := 350, CS := #CRNT_STEP, MST := "86_Times".STEP_MAX_TIME_STP_350, SC :=, BPFLT :=, AMST :=, FLT :=, ACT =>, DN =>)
      Contact( #STEP_350.DN )
      Move(in := 360, out1 => #CRNT_STEP)
   END_RUNG
   // the same network as SCL:
   #STEP_350(SN := 350, CS := #CRNT_STEP, MST := "86_Times".STEP_MAX_TIME_STP_350, ENO => #_w1);   // "500_SEQ_STEP"
   IF #_w1 AND #STEP_350.DN THEN #CRNT_STEP := 360; END_IF;
END_REGION

REGION Network 41: Step 360 = CV441 Closed Delay (Done = Jump To Step 410)
   RUNG wire#powerrail
      #STEP_360(SN := 360, CS := #CRNT_STEP, MST := "86_Times".STEP_MAX_TIME_STP_360, SC :=, BPFLT :=, AMST :=, FLT :=, ACT =>, DN =>)
      Contact( #STEP_360.DN )
      Move(in := 410, out1 => #CRNT_STEP)
   END_RUNG
   // the same network as SCL:
   #STEP_360(SN := 360, CS := #CRNT_STEP, MST := "86_Times".STEP_MAX_TIME_STP_360, ENO => #_w1);   // "500_SEQ_STEP"
   IF #_w1 AND #STEP_360.DN THEN #CRNT_STEP := 410; END_IF;
END_REGION

REGION Network 42: Step 370 = Close CV401
   RUNG wire#powerrail
      #STEP_370(SN := 370, CS := #CRNT_STEP, MST := "86_Times".STEP_MAX_TIME_STP_370, SC :=, BPFLT :=, AMST :=, FLT :=, ACT =>, DN =>)
      Contact( #STEP_370.DN )
      Move(in := 380, out1 => #CRNT_STEP)
   END_RUNG
   // the same network as SCL:
   #STEP_370(SN := 370, CS := #CRNT_STEP, MST := "86_Times".STEP_MAX_TIME_STP_370, ENO => #_w1);   // "500_SEQ_STEP"
   IF #_w1 AND #STEP_370.DN THEN #CRNT_STEP := 380; END_IF;
END_REGION

REGION Network 43: Step 380 = CV401 Closed Delay
